// TIA Portal project "XSFW_TIA31001_B0_V15.1" (V15.1) (continued)
END_REGION

REGION Network 63: Divider en marcha
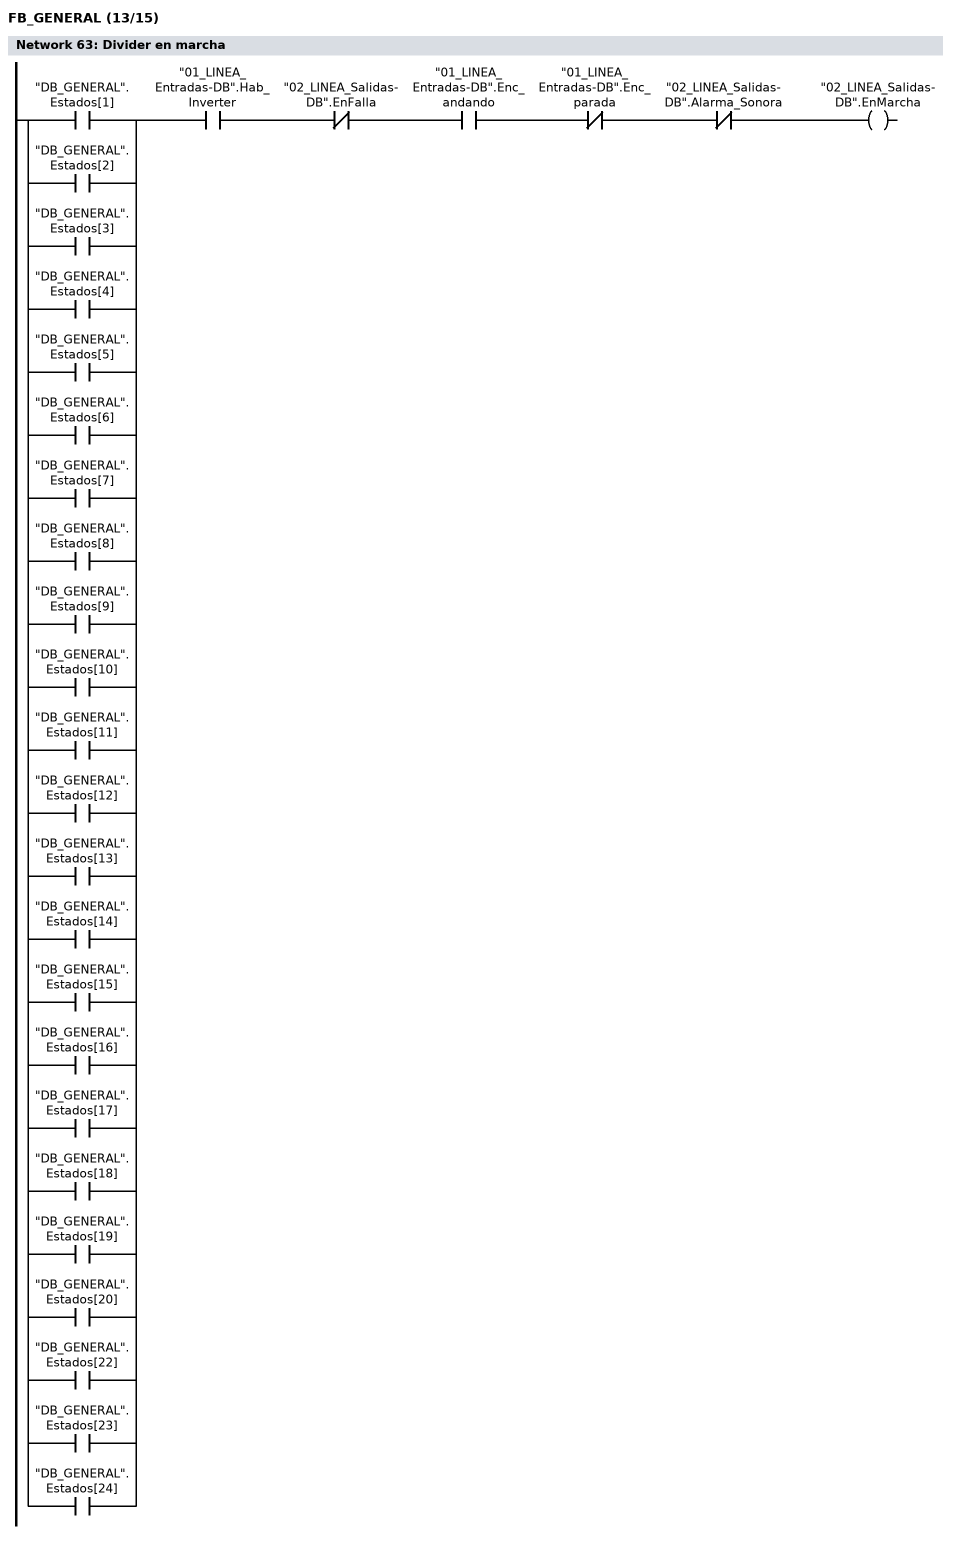
   RUNG wire#powerrail
      Contact( "DB_GENERAL".Estados[1] )
      wire#w1
      Contact( "01_LINEA_Entradas-DB".Hab_Inverter )
      I_Contact( "02_LINEA_Salidas-DB".EnFalla )
      Contact( "01_LINEA_Entradas-DB".Enc_andando )
      I_Contact( "01_LINEA_Entradas-DB".Enc_parada )
      I_Contact( "02_LINEA_Salidas-DB".Alarma_Sonora )
      Coil( "02_LINEA_Salidas-DB".EnMarcha )
   END_RUNG
   RUNG wire#powerrail
      Contact( "DB_GENERAL".Estados[2] )
   END_RUNG wire#w1
   RUNG wire#powerrail
      Contact( "DB_GENERAL".Estados[3] )
   END_RUNG wire#w1
   RUNG wire#powerrail
      Contact( "DB_GENERAL".Estados[4] )
   END_RUNG wire#w1
   RUNG wire#powerrail
      Contact( "DB_GENERAL".Estados[5] )
   END_RUNG wire#w1
   RUNG wire#powerrail
      Contact( "DB_GENERAL".Estados[6] )
   END_RUNG wire#w1
   RUNG wire#powerrail
      Contact( "DB_GENERAL".Estados[7] )
   END_RUNG wire#w1
   RUNG wire#powerrail
      Contact( "DB_GENERAL".Estados[8] )
   END_RUNG wire#w1
   RUNG wire#powerrail
      Contact( "DB_GENERAL".Estados[9] )
   END_RUNG wire#w1
   RUNG wire#powerrail
      Contact( "DB_GENERAL".Estados[10] )
   END_RUNG wire#w1
   RUNG wire#powerrail
      Contact( "DB_GENERAL".Estados[11] )
   END_RUNG wire#w1
   RUNG wire#powerrail
      Contact( "DB_GENERAL".Estados[12] )
   END_RUNG wire#w1
   RUNG wire#powerrail
      Contact( "DB_GENERAL".Estados[13] )
   END_RUNG wire#w1
   RUNG wire#powerrail
      Contact( "DB_GENERAL".Estados[14] )
   END_RUNG wire#w1
   RUNG wire#powerrail
      Contact( "DB_GENERAL".Estados[15] )
   END_RUNG wire#w1
   RUNG wire#powerrail
      Contact( "DB_GENERAL".Estados[16] )
   END_RUNG wire#w1
   RUNG wire#powerrail
      Contact( "DB_GENERAL".Estados[17] )
   END_RUNG wire#w1
   RUNG wire#powerrail
      Contact( "DB_GENERAL".Estados[18] )
   END_RUNG wire#w1
   RUNG wire#powerrail
      Contact( "DB_GENERAL".Estados[19] )
   END_RUNG wire#w1
   RUNG wire#powerrail
      Contact( "DB_GENERAL".Estados[20] )
   END_RUNG wire#w1
   RUNG wire#powerrail
      Contact( "DB_GENERAL".Estados[22] )
   END_RUNG wire#w1
   RUNG wire#powerrail
      Contact( "DB_GENERAL".Estados[23] )
   END_RUNG wire#w1
   RUNG wire#powerrail
      Contact( "DB_GENERAL".Estados[24] )
   END_RUNG wire#w1
   // the same network as SCL:
   "02_LINEA_Salidas-DB".EnMarcha := ("DB_GENERAL".Estados[1] OR "DB_GENERAL".Estados[2] OR "DB_GENERAL".Estados[3] OR "DB_GENERAL".Estados[4] OR "DB_GENERAL".Estados[5] OR "DB_GENERAL".Estados[6] OR "DB_GENERAL".Estados[7] OR "DB_GENERAL".Estados[8] OR "DB_GENERAL".Estados[9] OR "DB_GENERAL".Estados[10] OR "DB_GENERAL".Estados[11] OR "DB_GENERAL".Estados[12] OR "DB_GENERAL".Estados[13] OR "DB_GENERAL".Estados[14] OR "DB_GENERAL".Estados[15] OR "DB_GENERAL".Estados[16] OR "DB_GENERAL".Estados[17] OR "DB_GENERAL".Estados[18] OR "DB_GENERAL".Estados[19] OR "DB_GENERAL".Estados[20] OR "DB_GENERAL".Estados[22] OR "DB_GENERAL".Estados[23] OR "DB_GENERAL".Estados[24]) AND "01_LINEA_Entradas-DB".Hab_Inverter AND NOT "02_LINEA_Salidas-DB".EnFalla AND "01_LINEA_Entradas-DB".Enc_andando AND NOT "01_LINEA_Entradas-DB".Enc_parada AND NOT "02_LINEA_Salidas-DB".Alarma_Sonora;
END_REGION

REGION Network 64: Testigo de divider en marcha
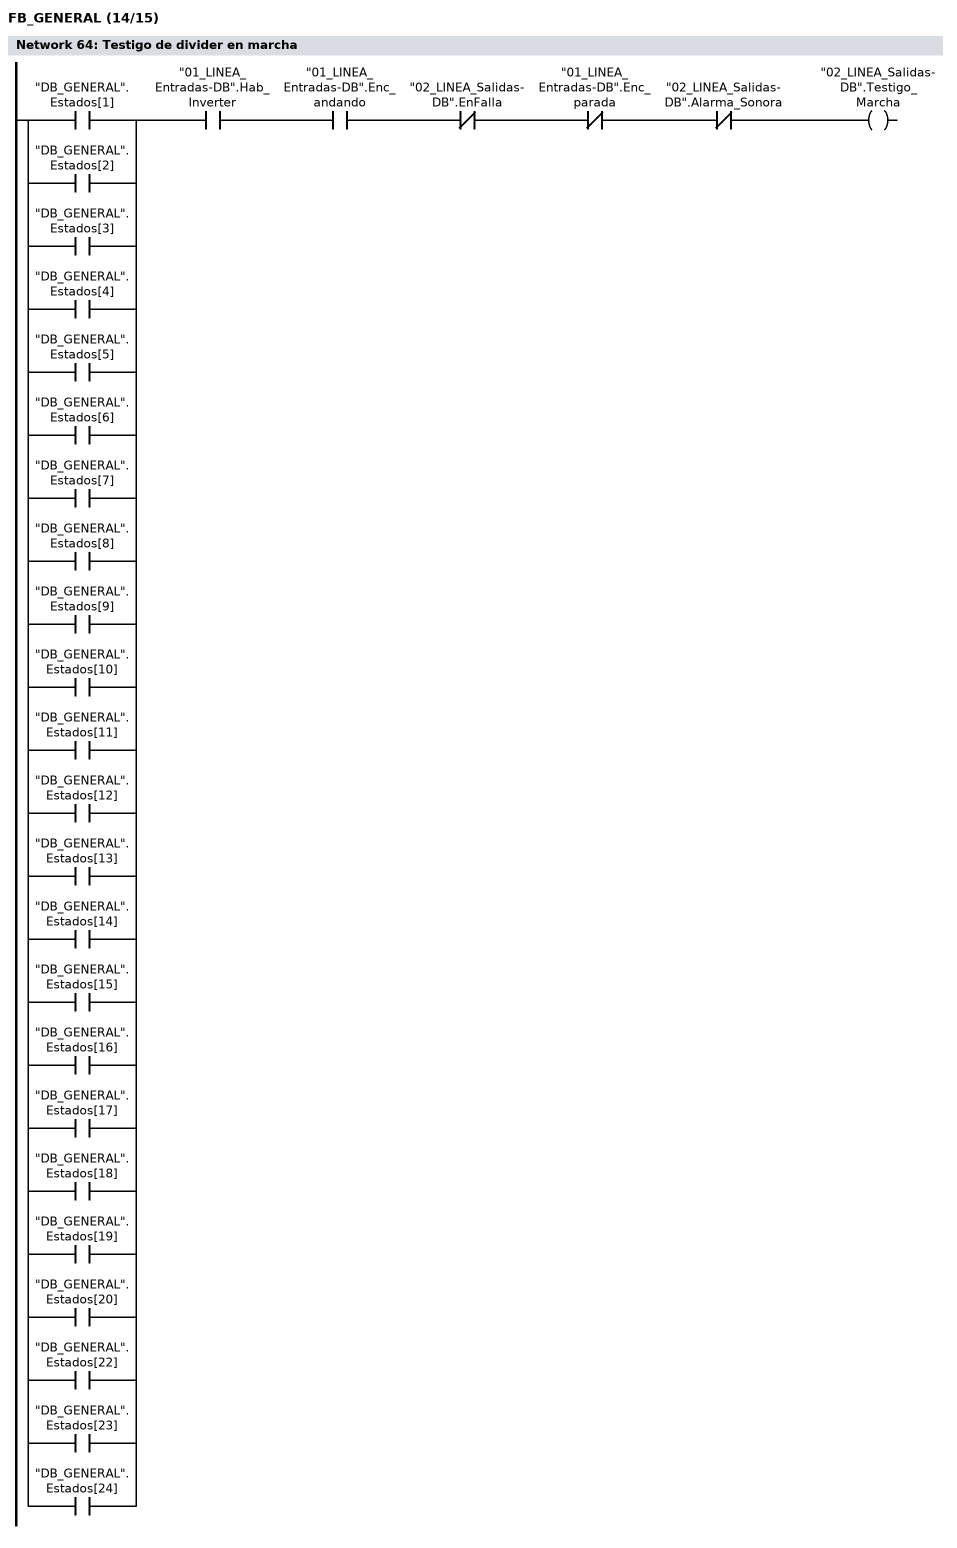
   RUNG wire#powerrail
      Contact( "DB_GENERAL".Estados[1] )
      wire#w1
      Contact( "01_LINEA_Entradas-DB".Hab_Inverter )
      Contact( "01_LINEA_Entradas-DB".Enc_andando )
      I_Contact( "02_LINEA_Salidas-DB".EnFalla )
      I_Contact( "01_LINEA_Entradas-DB".Enc_parada )
      I_Contact( "02_LINEA_Salidas-DB".Alarma_Sonora )
      Coil( "02_LINEA_Salidas-DB".Testigo_Marcha )
   END_RUNG
   RUNG wire#powerrail
      Contact( "DB_GENERAL".Estados[2] )
   END_RUNG wire#w1
   RUNG wire#powerrail
      Contact( "DB_GENERAL".Estados[3] )
   END_RUNG wire#w1
   RUNG wire#powerrail
      Contact( "DB_GENERAL".Estados[4] )
   END_RUNG wire#w1
   RUNG wire#powerrail
      Contact( "DB_GENERAL".Estados[5] )
   END_RUNG wire#w1
   RUNG wire#powerrail
      Contact( "DB_GENERAL".Estados[6] )
   END_RUNG wire#w1
   RUNG wire#powerrail
      Contact( "DB_GENERAL".Estados[7] )
   END_RUNG wire#w1
   RUNG wire#powerrail
      Contact( "DB_GENERAL".Estados[8] )
   END_RUNG wire#w1
   RUNG wire#powerrail
      Contact( "DB_GENERAL".Estados[9] )
   END_RUNG wire#w1
   RUNG wire#powerrail
      Contact( "DB_GENERAL".Estados[10] )
   END_RUNG wire#w1
   RUNG wire#powerrail
      Contact( "DB_GENERAL".Estados[11] )
   END_RUNG wire#w1
   RUNG wire#powerrail
      Contact( "DB_GENERAL".Estados[12] )
   END_RUNG wire#w1
   RUNG wire#powerrail
      Contact( "DB_GENERAL".Estados[13] )
   END_RUNG wire#w1
   RUNG wire#powerrail
      Contact( "DB_GENERAL".Estados[14] )
   END_RUNG wire#w1
   RUNG wire#powerrail
      Contact( "DB_GENERAL".Estados[15] )
   END_RUNG wire#w1
   RUNG wire#powerrail
      Contact( "DB_GENERAL".Estados[16] )
   END_RUNG wire#w1
   RUNG wire#powerrail
      Contact( "DB_GENERAL".Estados[17] )
   END_RUNG wire#w1
   RUNG wire#powerrail
      Contact( "DB_GENERAL".Estados[18] )
   END_RUNG wire#w1
   RUNG wire#powerrail
      Contact( "DB_GENERAL".Estados[19] )
   END_RUNG wire#w1
   RUNG wire#powerrail
      Contact( "DB_GENERAL".Estados[20] )
   END_RUNG wire#w1
   RUNG wire#powerrail
      Contact( "DB_GENERAL".Estados[22] )
   END_RUNG wire#w1
   RUNG wire#powerrail
      Contact( "DB_GENERAL".Estados[23] )
   END_RUNG wire#w1
   RUNG wire#powerrail
      Contact( "DB_GENERAL".Estados[24] )
   END_RUNG wire#w1
   // the same network as SCL:
   "02_LINEA_Salidas-DB".Testigo_Marcha := ("DB_GENERAL".Estados[1] OR "DB_GENERAL".Estados[2] OR "DB_GENERAL".Estados[3] OR "DB_GENERAL".Estados[4] OR "DB_GENERAL".Estados[5] OR "DB_GENERAL".Estados[6] OR "DB_GENERAL".Estados[7] OR "DB_GENERAL".Estados[8] OR "DB_GENERAL".Estados[9] OR "DB_GENERAL".Estados[10] OR "DB_GENERAL".Estados[11] OR "DB_GENERAL".Estados[12] OR "DB_GENERAL".Estados[13] OR "DB_GENERAL".Estados[14] OR "DB_GENERAL".Estados[15] OR "DB_GENERAL".Estados[16] OR "DB_GENERAL".Estados[17] OR "DB_GENERAL".Estados[18] OR "DB_GENERAL".Estados[19] OR "DB_GENERAL".Estados[20] OR "DB_GENERAL".Estados[22] OR "DB_GENERAL".Estados[23] OR "DB_GENERAL".Estados[24]) AND "01_LINEA_Entradas-DB".Hab_Inverter AND "01_LINEA_Entradas-DB".Enc_andando AND NOT "02_LINEA_Salidas-DB".EnFalla AND NOT "01_LINEA_Entradas-DB".Enc_parada AND NOT "02_LINEA_Salidas-DB".Alarma_Sonora;
END_REGION

REGION Network 65: Semaforo verde
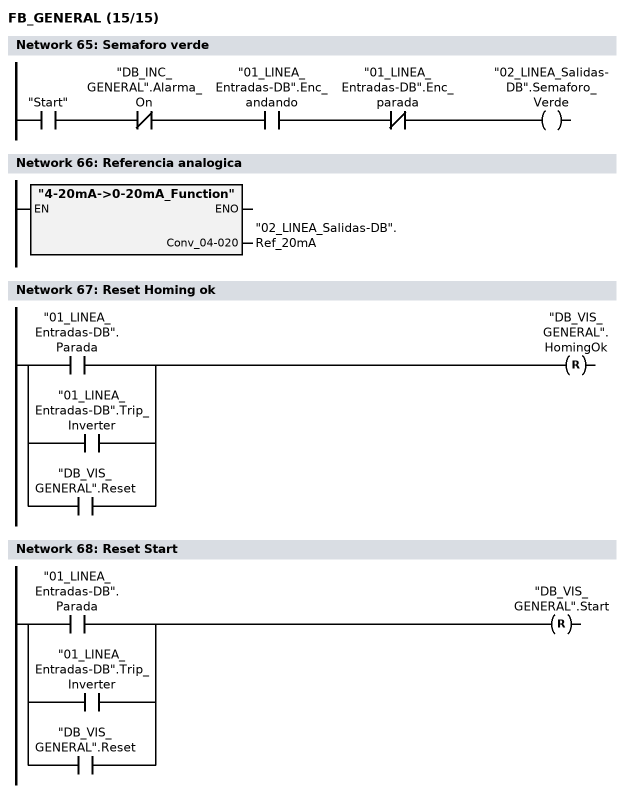
   RUNG wire#powerrail
      Contact( "Start" )
      I_Contact( "DB_INC_GENERAL".Alarma_On )
      Contact( "01_LINEA_Entradas-DB".Enc_andando )
      I_Contact( "01_LINEA_Entradas-DB".Enc_parada )
      Coil( "02_LINEA_Salidas-DB".Semaforo_Verde )
   END_RUNG
   // the same network as SCL:
   "02_LINEA_Salidas-DB".Semaforo_Verde := "Start" AND NOT "DB_INC_GENERAL".Alarma_On AND "01_LINEA_Entradas-DB".Enc_andando AND NOT "01_LINEA_Entradas-DB".Enc_parada;
END_REGION

REGION Network 66: Referencia analogica
   RUNG wire#powerrail
      "4-20mA->0-20mA_Function"("Conv_04-020" => "02_LINEA_Salidas-DB".Ref_20mA)
   END_RUNG
   // the same network as SCL:
   "4-20mA->0-20mA_Function"("Conv_04-020" => "02_LINEA_Salidas-DB".Ref_20mA);
END_REGION

REGION Network 67: Reset Homing ok
   RUNG wire#powerrail
      Contact( "01_LINEA_Entradas-DB".Parada )
      wire#w1
      R_Coil( "DB_VIS_GENERAL".HomingOk )
   END_RUNG
   RUNG wire#powerrail
      Contact( "01_LINEA_Entradas-DB".Trip_Inverter )
   END_RUNG wire#w1
   RUNG wire#powerrail
      Contact( "DB_VIS_GENERAL".Reset )
   END_RUNG wire#w1
   // the same network as SCL:
   IF "01_LINEA_Entradas-DB".Parada OR "01_LINEA_Entradas-DB".Trip_Inverter OR "DB_VIS_GENERAL".Reset THEN
       "DB_VIS_GENERAL".HomingOk := FALSE;
   END_IF;
END_REGION

REGION Network 68: Reset Start
   RUNG wire#powerrail
      Contact( "01_LINEA_Entradas-DB".Parada )
      wire#w1
      R_Coil( "DB_VIS_GENERAL".Start )
   END_RUNG
   RUNG wire#powerrail
      Contact( "01_LINEA_Entradas-DB".Trip_Inverter )
   END_RUNG wire#w1
   RUNG wire#powerrail
      Contact( "DB_VIS_GENERAL".Reset )
   END_RUNG wire#w1
   // the same network as SCL:
   IF "01_LINEA_Entradas-DB".Parada OR "01_LINEA_Entradas-DB".Trip_Inverter OR "DB_VIS_GENERAL".Reset THEN
       "DB_VIS_GENERAL".Start := FALSE;
   END_IF;
END_REGION
END_FUNCTION_BLOCK

FUNCTION "01_LINEA_Entradas" : Void   // FC1, LAD
TITLE = Bloque de entradas
{ S7_Optimized_Access := 'TRUE' }
VERSION : 0.1
BEGIN

REGION Network 1: Contador
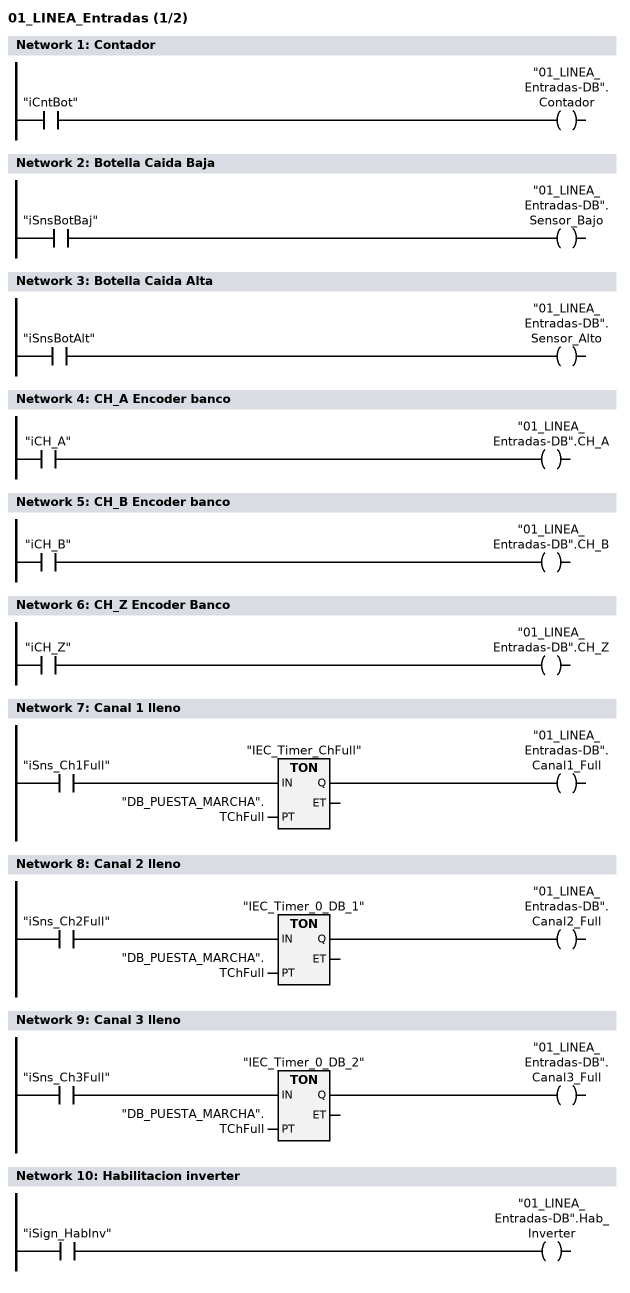
   RUNG wire#powerrail
      Contact( "iCntBot" )
      Coil( "01_LINEA_Entradas-DB".Contador )
   END_RUNG
   // the same network as SCL:
   "01_LINEA_Entradas-DB".Contador := "iCntBot";
END_REGION

REGION Network 2: Botella Caida Baja
   RUNG wire#powerrail
      Contact( "iSnsBotBaj" )
      Coil( "01_LINEA_Entradas-DB".Sensor_Bajo )
   END_RUNG
   // the same network as SCL:
   "01_LINEA_Entradas-DB".Sensor_Bajo := "iSnsBotBaj";
END_REGION

REGION Network 3: Botella Caida Alta
   RUNG wire#powerrail
      Contact( "iSnsBotAlt" )
      Coil( "01_LINEA_Entradas-DB".Sensor_Alto )
   END_RUNG
   // the same network as SCL:
   "01_LINEA_Entradas-DB".Sensor_Alto := "iSnsBotAlt";
END_REGION

REGION Network 4: CH_A Encoder banco
   RUNG wire#powerrail
      Contact( "iCH_A" )
      Coil( "01_LINEA_Entradas-DB".CH_A )
   END_RUNG
   // the same network as SCL:
   "01_LINEA_Entradas-DB".CH_A := "iCH_A";
END_REGION

REGION Network 5: CH_B Encoder banco
   RUNG wire#powerrail
      Contact( "iCH_B" )
      Coil( "01_LINEA_Entradas-DB".CH_B )
   END_RUNG
   // the same network as SCL:
   "01_LINEA_Entradas-DB".CH_B := "iCH_B";
END_REGION

REGION Network 6: CH_Z Encoder Banco
   RUNG wire#powerrail
      Contact( "iCH_Z" )
      Coil( "01_LINEA_Entradas-DB".CH_Z )
   END_RUNG
   // the same network as SCL:
   "01_LINEA_Entradas-DB".CH_Z := "iCH_Z";
END_REGION

REGION Network 7: Canal 1 lleno
   "IEC_Timer_ChFull".TON(IN := "iSns_Ch1Full", PT := "DB_PUESTA_MARCHA".TChFull);
   "01_LINEA_Entradas-DB".Canal1_Full := "IEC_Timer_ChFull".Q;
END_REGION

REGION Network 8: Canal 2 lleno
   "IEC_Timer_0_DB_1".TON(IN := "iSns_Ch2Full", PT := "DB_PUESTA_MARCHA".TChFull);
   "01_LINEA_Entradas-DB".Canal2_Full := "IEC_Timer_0_DB_1".Q;
END_REGION

REGION Network 9: Canal 3 lleno
   "IEC_Timer_0_DB_2".TON(IN := "iSns_Ch3Full", PT := "DB_PUESTA_MARCHA".TChFull);
   "01_LINEA_Entradas-DB".Canal3_Full := "IEC_Timer_0_DB_2".Q;
END_REGION

REGION Network 10: Habilitacion inverter
   RUNG wire#powerrail
      Contact( "iSign_HabInv" )
      Coil( "01_LINEA_Entradas-DB".Hab_Inverter )
   END_RUNG
   // the same network as SCL:
   "01_LINEA_Entradas-DB".Hab_Inverter := "iSign_HabInv";
END_REGION

REGION Network 11: Pulsador de Marcha de la columna 11
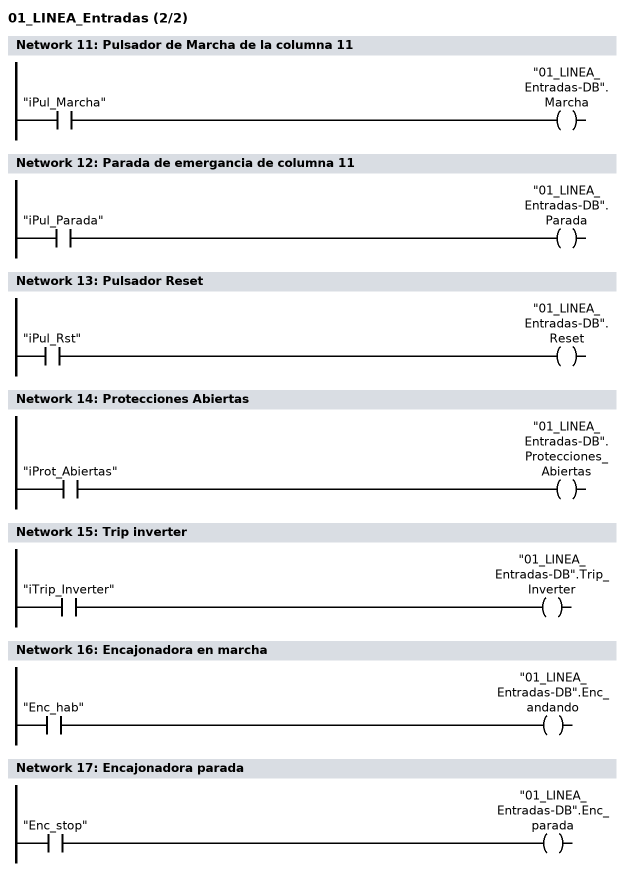
   RUNG wire#powerrail
      Contact( "iPul_Marcha" )
      Coil( "01_LINEA_Entradas-DB".Marcha )
   END_RUNG
   // the same network as SCL:
   "01_LINEA_Entradas-DB".Marcha := "iPul_Marcha";
END_REGION

REGION Network 12: Parada de emergancia de columna 11
   RUNG wire#powerrail
      Contact( "iPul_Parada" )
      Coil( "01_LINEA_Entradas-DB".Parada )
   END_RUNG
   // the same network as SCL:
   "01_LINEA_Entradas-DB".Parada := "iPul_Parada";
END_REGION

REGION Network 13: Pulsador Reset
   RUNG wire#powerrail
      Contact( "iPul_Rst" )
      Coil( "01_LINEA_Entradas-DB".Reset )
   END_RUNG
   // the same network as SCL:
   "01_LINEA_Entradas-DB".Reset := "iPul_Rst";
END_REGION

REGION Network 14: Protecciones Abiertas
   RUNG wire#powerrail
      Contact( "iProt_Abiertas" )
      Coil( "01_LINEA_Entradas-DB".Protecciones_Abiertas )
   END_RUNG
   // the same network as SCL:
   "01_LINEA_Entradas-DB".Protecciones_Abiertas := "iProt_Abiertas";
END_REGION

REGION Network 15: Trip inverter
   RUNG wire#powerrail
      Contact( "iTrip_Inverter" )
      Coil( "01_LINEA_Entradas-DB".Trip_Inverter )
   END_RUNG
   // the same network as SCL:
   "01_LINEA_Entradas-DB".Trip_Inverter := "iTrip_Inverter";
END_REGION

REGION Network 16: Encajonadora en marcha
   RUNG wire#powerrail
      Contact( "Enc_hab" )
      Coil( "01_LINEA_Entradas-DB".Enc_andando )
   END_RUNG
   // the same network as SCL:
   "01_LINEA_Entradas-DB".Enc_andando := "Enc_hab";
END_REGION

REGION Network 17: Encajonadora parada
   RUNG wire#powerrail
      Contact( "Enc_stop" )
      Coil( "01_LINEA_Entradas-DB".Enc_parada )
   END_RUNG
   // the same network as SCL:
   "01_LINEA_Entradas-DB".Enc_parada := "Enc_stop";
END_REGION
END_FUNCTION

FUNCTION "02_LINEA_Salidas" : Void   // FC2, LAD
{ S7_Optimized_Access := 'TRUE' }
VERSION : 0.1
BEGIN

REGION Network 1: Alarma Sonora
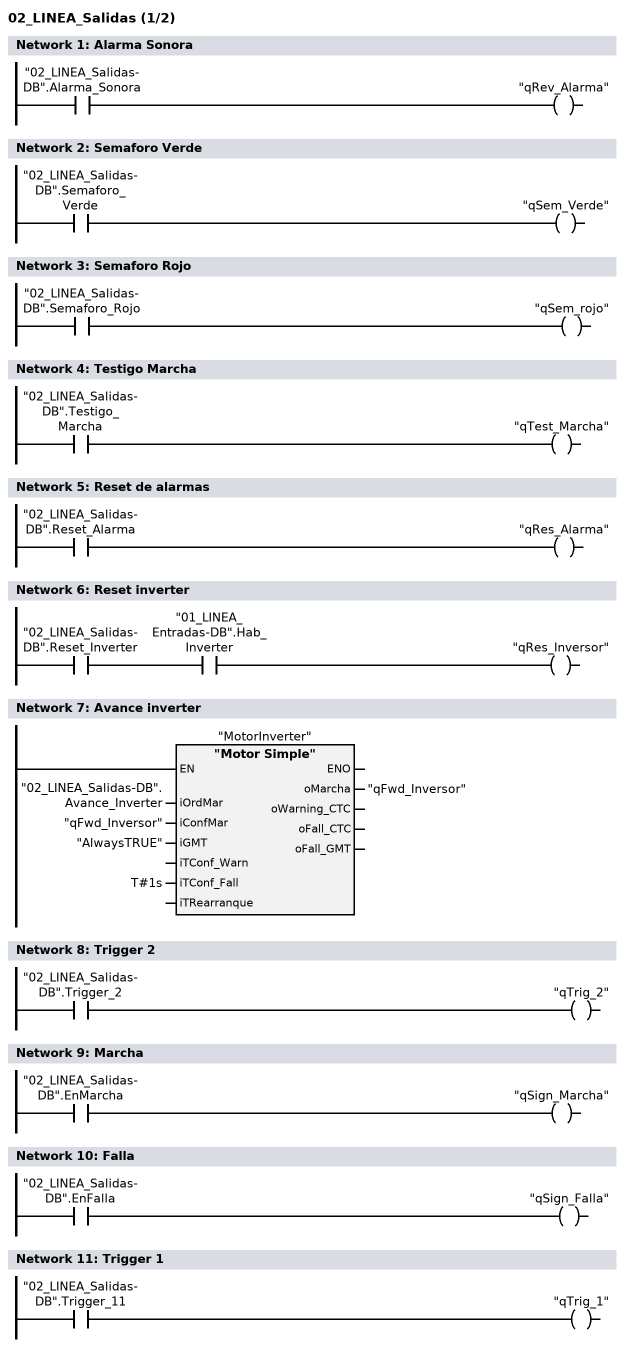
   RUNG wire#powerrail
      Contact( "02_LINEA_Salidas-DB".Alarma_Sonora )
      Coil( "qRev_Alarma" )
   END_RUNG
   // the same network as SCL:
   "qRev_Alarma" := "02_LINEA_Salidas-DB".Alarma_Sonora;
END_REGION

REGION Network 2: Semaforo Verde
   RUNG wire#powerrail
      Contact( "02_LINEA_Salidas-DB".Semaforo_Verde )
      Coil( "qSem_Verde" )
   END_RUNG
   // the same network as SCL:
   "qSem_Verde" := "02_LINEA_Salidas-DB".Semaforo_Verde;
END_REGION

REGION Network 3: Semaforo Rojo
   RUNG wire#powerrail
      Contact( "02_LINEA_Salidas-DB".Semaforo_Rojo )
      Coil( "qSem_rojo" )
   END_RUNG
   // the same network as SCL:
   "qSem_rojo" := "02_LINEA_Salidas-DB".Semaforo_Rojo;
END_REGION

REGION Network 4: Testigo Marcha
   RUNG wire#powerrail
      Contact( "02_LINEA_Salidas-DB".Testigo_Marcha )
      Coil( "qTest_Marcha" )
   END_RUNG
   // the same network as SCL:
   "qTest_Marcha" := "02_LINEA_Salidas-DB".Testigo_Marcha;
END_REGION

REGION Network 5: Reset de alarmas
   RUNG wire#powerrail
      Contact( "02_LINEA_Salidas-DB".Reset_Alarma )
      Coil( "qRes_Alarma" )
   END_RUNG
   // the same network as SCL:
   "qRes_Alarma" := "02_LINEA_Salidas-DB".Reset_Alarma;
END_REGION

REGION Network 6: Reset inverter
   RUNG wire#powerrail
      Contact( "02_LINEA_Salidas-DB".Reset_Inverter )
      Contact( "01_LINEA_Entradas-DB".Hab_Inverter )
      Coil( "qRes_Inversor" )
   END_RUNG
   // the same network as SCL:
   "qRes_Inversor" := "02_LINEA_Salidas-DB".Reset_Inverter AND "01_LINEA_Entradas-DB".Hab_Inverter;
END_REGION

REGION Network 7: Avance inverter
   RUNG wire#powerrail
      "MotorInverter"(iOrdMar := "02_LINEA_Salidas-DB".Avance_Inverter, iConfMar := "qFwd_Inversor", iGMT := "AlwaysTRUE", iTConf_Warn :=, iTConf_Fall := T#1s, iTRearranque :=, oMarcha => "qFwd_Inversor", oWarning_CTC =>, oFall_CTC =>, oFall_GMT =>)
   END_RUNG
   // the same network as SCL:
   "MotorInverter"(iOrdMar := "02_LINEA_Salidas-DB".Avance_Inverter,   // "Motor Simple"
                   iConfMar := "qFwd_Inversor",
                   iGMT := "AlwaysTRUE",
                   iTConf_Fall := T#1s,
                   oMarcha => "qFwd_Inversor");
END_REGION

REGION Network 8: Trigger 2
   RUNG wire#powerrail
      Contact( "02_LINEA_Salidas-DB".Trigger_2 )
      Coil( "qTrig_2" )
   END_RUNG
   // the same network as SCL:
   "qTrig_2" := "02_LINEA_Salidas-DB".Trigger_2;
END_REGION

REGION Network 9: Marcha
   RUNG wire#powerrail
      Contact( "02_LINEA_Salidas-DB".EnMarcha )
      Coil( "qSign_Marcha" )
   END_RUNG
   // the same network as SCL:
   "qSign_Marcha" := "02_LINEA_Salidas-DB".EnMarcha;
END_REGION

REGION Network 10: Falla
   RUNG wire#powerrail
      Contact( "02_LINEA_Salidas-DB".EnFalla )
      Coil( "qSign_Falla" )
   END_RUNG
   // the same network as SCL:
   "qSign_Falla" := "02_LINEA_Salidas-DB".EnFalla;
END_REGION

REGION Network 11: Trigger 1
   RUNG wire#powerrail
      Contact( "02_LINEA_Salidas-DB".Trigger_11 )
      Coil( "qTrig_1" )
   END_RUNG
   // the same network as SCL:
   "qTrig_1" := "02_LINEA_Salidas-DB".Trigger_11;
END_REGION

REGION Network 12: Trigger 22
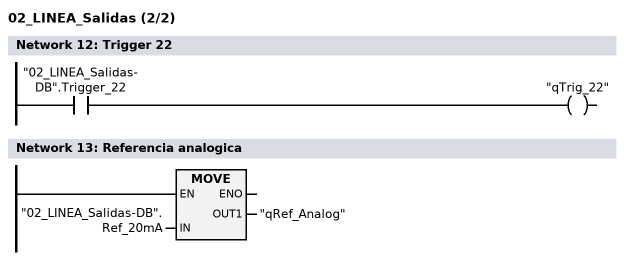
   RUNG wire#powerrail
      Contact( "02_LINEA_Salidas-DB".Trigger_22 )
      Coil( "qTrig_22" )
   END_RUNG
   // the same network as SCL:
   "qTrig_22" := "02_LINEA_Salidas-DB".Trigger_22;
END_REGION

REGION Network 13: Referencia analogica
   RUNG wire#powerrail
      Move(in := "02_LINEA_Salidas-DB".Ref_20mA, out1 => "qRef_Analog")
   END_RUNG
   // the same network as SCL:
   "qRef_Analog" := "02_LINEA_Salidas-DB".Ref_20mA;
END_REGION
END_FUNCTION

FUNCTION "4-20mA->0-20mA_Function" : Void   // FC3, LAD
TITLE = Conversion 4-20 -> 0-20 Canal 1
{ S7_Optimized_Access := 'TRUE' }
VERSION : 0.1
   VAR_OUTPUT
      "Conv_04-020" : Int;
   END_VAR
   VAR_TEMP
      Input_Analog1 : Real;
      Temp_Analog1 : Real;
      Input_Analog2 : Real;
      Temp_Analog2 : Real;
   END_VAR
BEGIN

REGION Network 1
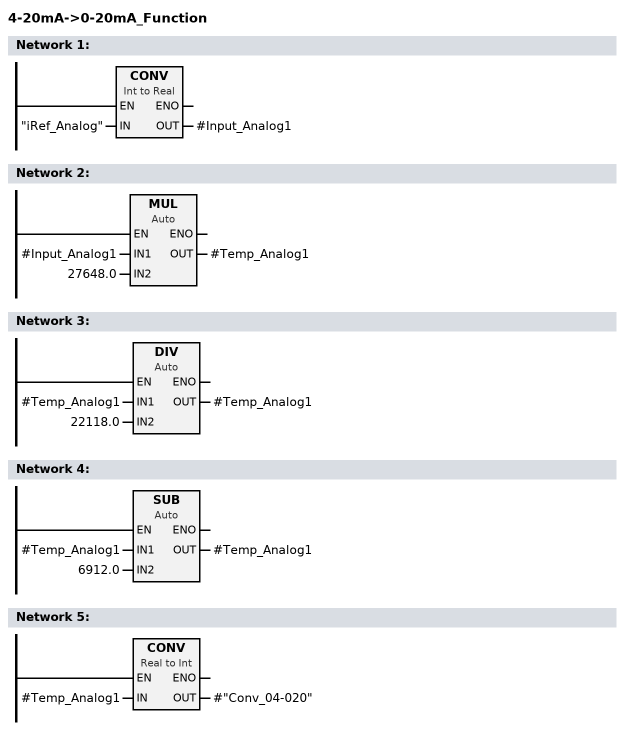
   RUNG wire#powerrail
      { S7_Templates := "[SrcType := Int, DestType := Real]" } Convert(in := "iRef_Analog", out => #Input_Analog1)
   END_RUNG
   // the same network as SCL:
   #Input_Analog1 := INT_TO_REAL("iRef_Analog");
END_REGION

REGION Network 2
   RUNG wire#powerrail
      Mul(in1 := #Input_Analog1, in2 := 27648.0, out => #Temp_Analog1)
   END_RUNG
   // the same network as SCL:
   #Temp_Analog1 := #Input_Analog1 * 27648.0;
END_REGION

REGION Network 3
   RUNG wire#powerrail
      Div(in1 := #Temp_Analog1, in2 := 22118.0, out => #Temp_Analog1)
   END_RUNG
   // the same network as SCL:
   #Temp_Analog1 := #Temp_Analog1 / 22118.0;
END_REGION

REGION Network 4
   RUNG wire#powerrail
      Sub(in1 := #Temp_Analog1, in2 := 6912.0, out => #Temp_Analog1)
   END_RUNG
   // the same network as SCL:
   #Temp_Analog1 := #Temp_Analog1 - 6912.0;
END_REGION

REGION Network 5
   RUNG wire#powerrail
      { S7_Templates := "[SrcType := Real, DestType := Int]" } Convert(in := #Temp_Analog1, out => #"Conv_04-020")
   END_RUNG
   // the same network as SCL:
   #"Conv_04-020" := REAL_TO_INT(#Temp_Analog1);
END_REGION
END_FUNCTION

ORGANIZATION_BLOCK "Main"   // OB1, LAD, ProgramCycle
TITLE = "Main Program Sweep (Cycle)"
{ S7_Optimized_Access := 'TRUE' }
VERSION : 0.1
   VAR_INPUT
      Initial_Call : Bool;   // Initial call of this OB
      Remanence : Bool;   // =True, if remanent data are available
   END_VAR
BEGIN

REGION Network 1: Asigno entradas a variables
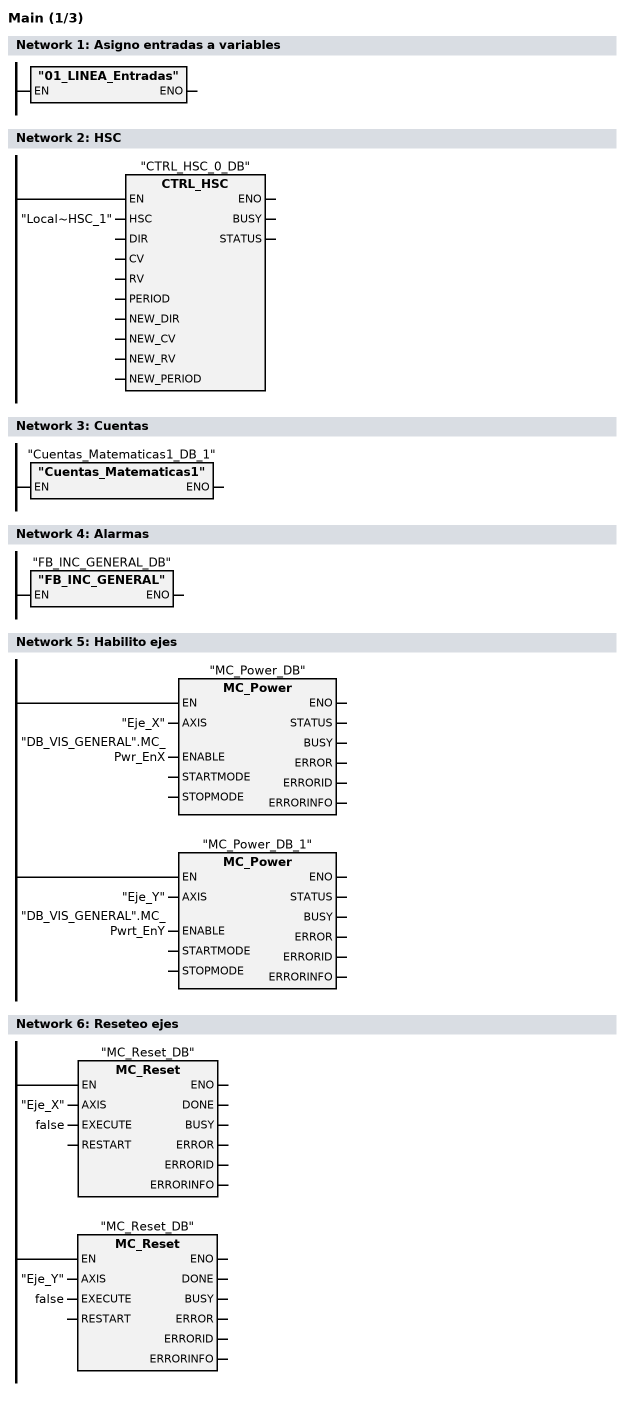
   RUNG wire#powerrail
      "01_LINEA_Entradas"()
   END_RUNG
   // the same network as SCL:
   "01_LINEA_Entradas"();
END_REGION

REGION Network 2: HSC
   "CTRL_HSC_0_DB"(HSC := "Local~HSC_1");   // CTRL_HSC
END_REGION

REGION Network 3: Cuentas
   RUNG wire#powerrail
      "Cuentas_Matematicas1_DB_1"()
   END_RUNG
   // the same network as SCL:
   "Cuentas_Matematicas1_DB_1"();   // "Cuentas_Matematicas1"
END_REGION

REGION Network 4: Alarmas
   RUNG wire#powerrail
      "FB_INC_GENERAL_DB"()
   END_RUNG
   // the same network as SCL:
   "FB_INC_GENERAL_DB"();   // "FB_INC_GENERAL"
END_REGION

REGION Network 5: Habilito ejes
   "MC_Power_DB"(Axis := "Eje_X", Enable := "DB_VIS_GENERAL".MC_Pwr_EnX);   // MC_Power
   "MC_Power_DB_1"(Axis := "Eje_Y", Enable := "DB_VIS_GENERAL".MC_Pwrt_EnY);   // MC_Power
END_REGION

REGION Network 6: Reseteo ejes
   "MC_Reset_DB"(Axis := "Eje_X", Execute := false);   // MC_Reset
   "MC_Reset_DB"(Axis := "Eje_Y", Execute := false);   // MC_Reset
END_REGION

REGION Network 7: Llamo a FB General
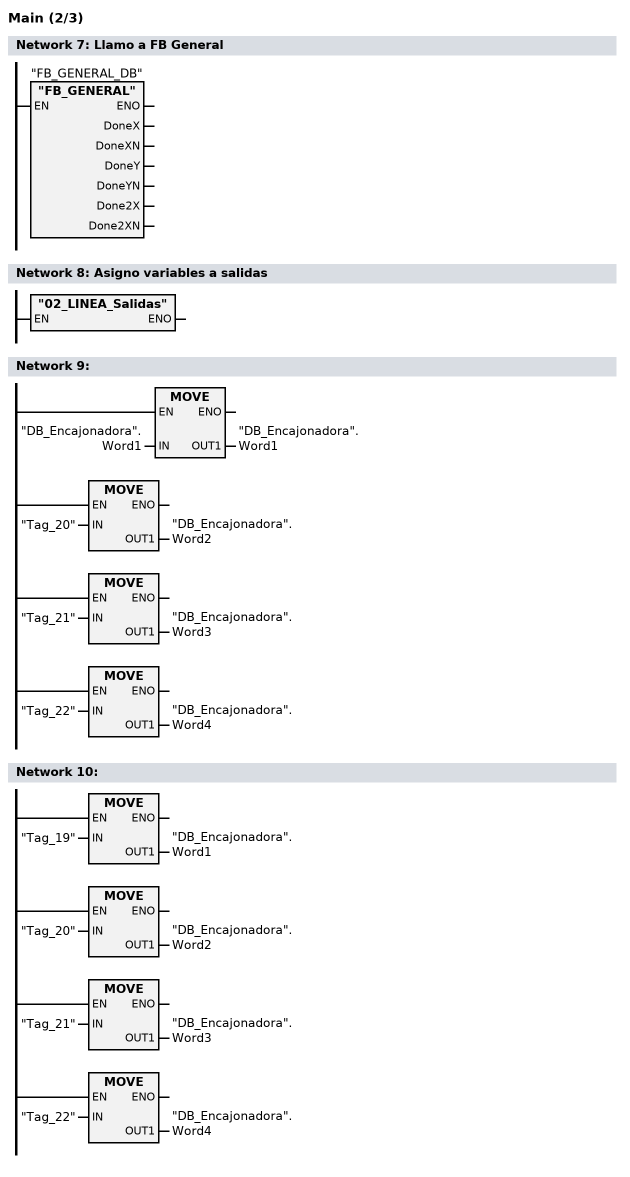
   RUNG wire#powerrail
      "FB_GENERAL_DB"(DoneX =>, DoneY =>, Done2X =>, DoneXN =>, DoneYN =>, Done2XN =>)
   END_RUNG
   // the same network as SCL:
   "FB_GENERAL_DB"();   // "FB_GENERAL"
END_REGION

REGION Network 8: Asigno variables a salidas
   RUNG wire#powerrail
      "02_LINEA_Salidas"()
   END_RUNG
   // the same network as SCL:
   "02_LINEA_Salidas"();
END_REGION

REGION Network 9
   RUNG wire#powerrail
      Move(in := "DB_Encajonadora".Word1, out1 => "DB_Encajonadora".Word1)
   END_RUNG
   RUNG wire#powerrail
      Move(in := "Tag_20", out1 => "DB_Encajonadora".Word2)
   END_RUNG
   RUNG wire#powerrail
      Move(in := "Tag_21", out1 => "DB_Encajonadora".Word3)
   END_RUNG
   RUNG wire#powerrail
      Move(in := "Tag_22", out1 => "DB_Encajonadora".Word4)
   END_RUNG
   // the same network as SCL:
   "DB_Encajonadora".Word1 := "DB_Encajonadora".Word1;
   "DB_Encajonadora".Word2 := "Tag_20";
   "DB_Encajonadora".Word3 := "Tag_21";
   "DB_Encajonadora".Word4 := "Tag_22";
END_REGION

REGION Network 10
   RUNG wire#powerrail
      Move(in := "Tag_19", out1 => "DB_Encajonadora".Word1)
   END_RUNG
   RUNG wire#powerrail
      Move(in := "Tag_20", out1 => "DB_Encajonadora".Word2)
   END_RUNG
   RUNG wire#powerrail
      Move(in := "Tag_21", out1 => "DB_Encajonadora".Word3)
   END_RUNG
   RUNG wire#powerrail
      Move(in := "Tag_22", out1 => "DB_Encajonadora".Word4)
   END_RUNG
   // the same network as SCL:
   "DB_Encajonadora".Word1 := "Tag_19";
   "DB_Encajonadora".Word2 := "Tag_20";
   "DB_Encajonadora".Word3 := "Tag_21";
   "DB_Encajonadora".Word4 := "Tag_22";
END_REGION

REGION Network 11
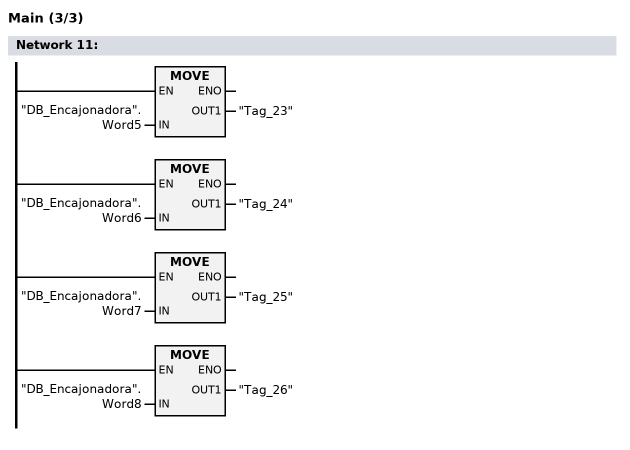
   RUNG wire#powerrail
      Move(in := "DB_Encajonadora".Word5, out1 => "Tag_23")
   END_RUNG
   RUNG wire#powerrail
      Move(in := "DB_Encajonadora".Word6, out1 => "Tag_24")
   END_RUNG
   RUNG wire#powerrail
      Move(in := "DB_Encajonadora".Word7, out1 => "Tag_25")
   END_RUNG
   RUNG wire#powerrail
      Move(in := "DB_Encajonadora".Word8, out1 => "Tag_26")
   END_RUNG
   // the same network as SCL:
   "Tag_23" := "DB_Encajonadora".Word5;
   "Tag_24" := "DB_Encajonadora".Word6;
   "Tag_25" := "DB_Encajonadora".Word7;
   "Tag_26" := "DB_Encajonadora".Word8;
END_REGION
END_ORGANIZATION_BLOCK

ORGANIZATION_BLOCK "Cyclic interrupt"   // OB30, LAD, CyclicInterrupt
{ S7_Optimized_Access := 'TRUE' }
VERSION : 0.1
   VAR_INPUT
      Initial_Call : Bool;   // Initial call of this OB
      Event_Count : Int;   // Events discarded
   END_VAR
BEGIN

REGION Network 1: Move
